VERSION : 0.1
// Data area for commands from master PLC
   VAR
      CRNT_MODE : Int := 1;   // 1 = Auto, 2 = Man, 3 = FatAuto, 4 = FatMan
      HEART_BEAT : Bool;   // Heartbeat
      ESTOP_OK : Bool;   // 1 = OK, 0 = Estop active
      RST_AUT_SEQ : Bool;   // Reset automatic sequence
      RUN_E131 : Bool;   // IA Compressor demand
      RUN_P301 : Bool;   // 1 = Run, 0 = Not
      RUN_BC_SEQ : Bool;   // 1 = Start command. 0 = Not
      PB_STS_CNFMD : Bool;   // Pilot burn status confirmed by IGG
      CRG_BLNK_MODE : Bool;   // 1 = Cargon blanketing mode, 0 = Not
      RUN_BC_O2_RAMP : Bool;   // 1 = Run ramp, 0 = Not
      BC_SD_CMND : Bool;   // 1 = Run. 0 = Shutdown
      STOP_BURNS_CMND : Bool;   // 1 = Burners off, 0 = Not
      CLS_CV127_CMND : Bool;   // 1 = OPEN, 0 = Close
      CLS_CV203_CMND : Bool;   // 1 = Close, 0 = Not
      CLS_CV111_CMND : Bool;   // 1 = Close, 0 = Not
      IGG_ALARM : Bool;   // 1 = IGG Alarm state, 0 = Not
      RUN_P305 : Bool;   // Fresh water pump demand
      CV403_OPEN : Bool;   // 1 = Valve is open, 0 = Not
      "E 500A RUN" : Bool;   // Fuel Pump 1 Enabled
      "E 500B RUN" : Bool;   // Fuel Pump 2 Enabled
      "TIT 360 Healthy" : Bool;   // Outlet CSW Temp TIT360
      "TIT 401 Healthy" : Bool;   // IG Temp
      "PIT 316 Healthy" : Bool;   // Outlet CSW Pressure
      RST_LOCKOUT : Bool;   // Reset alarms
      "CA Blower Running" : Bool;   // E139-MCCP/6TA1
      Alarm_Reset : Bool;   // Alarm_Reset
      BWT_MODE : Bool;
      "P301 PRSNT" : Bool;
      "TIT 315 Healthy" : Bool;   // PIT 315 Healthy
      SFTY_SYS_IL : Bool;   // SFTY_SYS_IL
      "Master Stop" : Bool;   // Master Stop
      "CV401 Closed" : Bool;   // CV401 Closed
      SPR_5_7 : Bool;   // Spare bool
      IGG_CRNT_STEP : Int;   // IGG Current Step
   END_VAR
BEGIN
END_DATA_BLOCK

DATA_BLOCK "55_STATUS_DATA"   // DB55
TITLE = Status Data
{ S7_Optimized_Access := 'FALSE' }
AUTHOR : JRS
VERSION : 0.1
// Data area for status to master PLC
   VAR
      PIT112_SCALED : Real;   // IA Inlet pressure
      CV203_CNTRL : Real;   // Main fuel reg Valve Control
      PIT204_SCALED : Real;   // IGG Inlet fuel pressure
      CRNT_MODE : Int := 1;   // 1 = Auto, 2 = Man, 3 = FatAuto, 4 = FatMan
      HEART_BEAT : Bool;   // Heartbeat
      AUT_SEQ_RNG : Bool;   // Auto sequence running
      VLVS_AT_INIT : Bool;   // All valves in initial state
      P301_ENBLD : Bool;   // P301 enabled input sent from BC
      P301_TRIPPED : Bool;   // P301 tripped input sent from BC
      TS006_OK : Bool;   // TS006 Is healthy
      TS403_OK : Bool;   // TS403 Is healthy
      LS001_OK : Bool;   // LS001 Is healthy
      E131_RUNNING : Bool;   // E131 Running
      BC_SEQ_STARTED : Bool;   // BC Sequence confirmed as started
      PILOT_BURNER_ACTV : Bool;   // Pilot burn confirmed as active
      PILOT_PURGE_DN : Bool;   // Pilot burner purge completed
      RAMPING_O2_ACTV : Bool;   // Ramping of O2 is active
      O2_LVL_OK : Bool;   // O2 Level within specification
      SHTNG_DN_CNF : Bool;   // Shutting down confirmed
      O2_CNTRL_STPD : Bool;   // O2 Control modulation stopped
      BURNS_STOPPED : Bool;   // Confirmation burners are off
      CV127_CLOSED : Bool;   // CV127 Closed status
      CV203_CLOSED : Bool;   // CV203 Closed status
      CV111_CLOSED : Bool;   // CV111 Closed status
      BC_SD_DONE : Bool;   // BC Shutdown sequence done
      BC_ALARM : Bool;   // 1 = BC Alarm state, 0 = Not
      MAA_PRES_IN_RNG : Bool;   // PIT113 Main atom air pressure within range
      "FD001FDU Healthy" : Bool;   // FDU Healthy
      "FS 317 Healthy" : Bool;   // Jacket Cooling Water Flow Switch
      "PIT 204 Healthy" : Bool;   // PIT 204 Healthy
      "FS 320 Healthy" : Bool;   // FS 320 Healthy
      Warnings : Bool;   // Warnings
      "PIT 112 Healthy" : Bool;   // PIT 112 Healthy
      MAIN_BURNER_ACTV : Bool;   // MAIN_BURNER_ACTV
      "BC New ALARM" : Bool;   // New alarm
      "BC New WARNING" : Bool;   // New warning
      P305_ENBLD : Bool;   // P305 enabled input sent from BC
      P305_TRIPPED : Bool;   // P305 tripped input sent from BC
      P305_PRSNT : Bool;   // P305_PRSNT
      SPR_18_3 : Bool;   // Spare bit
      SPR_18_4 : Bool;   // Spare bit
      SPR_18_5 : Bool;   // Spare bit
      SPR_18_6 : Bool;   // Spare bit
      SPR_18_7 : Bool;   // Spare bit
   END_VAR
BEGIN
END_DATA_BLOCK

DATA_BLOCK "57_COMMS_DATE_TIME"   // DB57
{ S7_Optimized_Access := 'FALSE' }
VERSION : 0.1
   VAR
      SYSTEM_TIME : DTL;
      LOCAL_TIME : DTL;
   END_VAR
BEGIN
END_DATA_BLOCK

DATA_BLOCK "59_COMMS_HEALTH_DATA"   // DB59
TITLE = Communications Health Data
{ S7_Optimized_Access := 'TRUE' }
AUTHOR : JRS
VERSION : 0.1
// Data area for communications health determination
   VAR
      CLOCK_POS_EDGE : Bool;   // Edge bit
      CLOCK_NEG_EDGE : Bool;   // Edge bit
      MSTR_TRUE_TMR : TON_TIME;
      MSTR_FALSE_TMR : TON_TIME;
      MSTR_HB_MISSING : Bool;   // Heatbeat missing flag
   END_VAR
BEGIN
   MSTR_FALSE_TMR.PT := T#2s;
   MSTR_TRUE_TMR.PT := T#2s;
END_DATA_BLOCK

// folder: 60 - 69 Alarm & Satus Handling

DATA_BLOCK "60_Alarm_Data"   // DB60
{ S7_Optimized_Access := 'FALSE' }
VERSION : 0.1
   VAR
      BC_ALARM_WORD_01 : Word;
      BC_ALARM_WORD_02 : Word;
      BC_ALARM_WORD_03 : Word;
      BC_ALARM_WORD_04 : Word;
      BC_ALARM_WORD_05 : Word;
      BC_ALARM_WORD_06 : Word;
      BC_ALARM_WORD_07 : Word;
      BC_ALARM_WORD_08 : Word;
      BC_ALARM_WORD_09 : Word;
      BC_ALARM_WORD_10 : Word;
      BC_ALARM_WORD_11 : Word;
      BC_ALARM_WORD_12 : Word;
      BC_ALARM_WORD_13 : Word;
      BC_ALARM_WORD_14 : Word;
      BC_ALARM_WORD_15 : Word;
      BC_ALARM_WORD_16 : Word;
      ALRM_PRSNT : Bool;
   END_VAR
BEGIN
END_DATA_BLOCK

DATA_BLOCK "62_Warning_Data"   // DB62
{ S7_Optimized_Access := 'FALSE' }
VERSION : 0.1
   VAR
      BC_WARNING_WORD_01 : Word;   // PIT 204
      BC_WARNING_WORD_02 : Word;   // TIT 202
      BC_WARNING_WORD_03 : Word;   // PIT 205
      BC_WARNING_WORD_04 : Word;   // PIT 112
      BC_WARNING_WORD_05 : Word;   // PIT 113
      BC_WARNING_WORD_06 : Word;
      BC_WARNING_WORD_07 : Word;
      BC_WARNING_WORD_08 : Word;
      WRNG_PRSNT : Bool;
   END_VAR
BEGIN
END_DATA_BLOCK

DATA_BLOCK "503_WARNING CHCK_DB"   // DB63
{ S7_Optimized_Access := 'TRUE' }
VERSION : 0.1
// stored: InstanceOfName 503_ALARM CHCK
"503_ALARM CHCK"
BEGIN
END_DATA_BLOCK

DATA_BLOCK "64_Message_Data"   // DB64
{ S7_Optimized_Access := 'FALSE' }
VERSION : 0.1
   VAR
      BC_MESSAGE_WORD_01 : Word;
      BC_MESSAGE_WORD_02 : Word;
      BC_MESSAGE_WORD_03 : Word;
      BC_MESSAGE_WORD_04 : Word;
      BC_MESSAGE_WORD_05 : Word;
      BC_MESSAGE_WORD_06 : Word;
      BC_MESSAGE_WORD_07 : Word;
      BC_MESSAGE_WORD_08 : Word;
      MSG_PRSNT : Bool;
   END_VAR
BEGIN
END_DATA_BLOCK

DATA_BLOCK "503_ALARM CHCK_DB"   // DB65
{ S7_Optimized_Access := 'TRUE' }
VERSION : 0.1
// stored: InstanceOfName 503_ALARM CHCK
"503_ALARM CHCK"
BEGIN
END_DATA_BLOCK

DATA_BLOCK "66_Event_Data"   // DB66
{ S7_Optimized_Access := 'FALSE' }
VERSION : 0.1
   VAR
      BC_EVENT_WORD_01 : Word;
      BC_EVENT_WORD_02 : Word;
      BC_EVENT_WORD_03 : Word;
      BC_EVENT_WORD_04 : Word;
      BC_EVENT_WORD_05 : Word;
      BC_EVENT_WORD_06 : Word;
      BC_EVENT_WORD_07 : Word;
      BC_EVENT_WORD_08 : Word;
      EVENT_PRSNT : Bool;
   END_VAR
BEGIN
END_DATA_BLOCK

DATA_BLOCK "68_Sys_Status_Data"   // DB68
TITLE = System Status Data
{ S7_Optimized_Access := 'TRUE' }
AUTHOR : JRS
VERSION : 0.1
// Data area for system status information as required by the code
   VAR
      VLVS_AT_INIT : Bool;   // All valves at initial position
      INTRLKS_OK : Bool;   // System interlocks ok
      IA_PRES_IN_RNG : Bool;   // IA Pressure Within Range - PIT112
      CSW_IL_PRES_IN_RNG : Bool;   // CSW Inlet pressure within range - PIT359
      FUEL_PRES_IN_RNG : Bool;   // Fuel pressure within range - PIT204
      OP_PRES_IN_RNG : Bool;   // Output pressure within range - PIT402
      VALID_FLAME : Bool;   // Flame detection & > min value - FD001
      O2_INTO_SPEC_DLY : TON_TIME;   // O2 Going into specification de-bounce timer
      O2_OUT_SPEC_DLY : TOF_TIME;   // O2 Going out of specification de-bounce timer
      O2_WITHIN_SPEC : Bool;   // O2 Contenct is within specification
      SHT_DN_CNF_DLY : TP_TIME;   // Shutting down confirmed timer
      O2_CNTRL_STPPD_DLY : TP_TIME;   // O2 Control stopped confirmed timer
      BURNS_STPPD_DLY : TP_TIME;   // Burns stopped confirmed timer
      CV127_CLSD_DLY : TP_TIME;   // CV127 Closed confirmed timer
      CV203_CLSD_DLY : TON_TIME;   // CV203 Closed confirmed timer
      CV111_CLSD_DLY : TON_TIME;   // CV111 Closed confirmed timer
      BC_SD_DONE : TP_TIME;   // BC Shutdown done timer
      CV127_CLSD_FLG : Bool;
   END_VAR
BEGIN
END_DATA_BLOCK

DATA_BLOCK "Main Burner Animation_DB"   // DB69
{ S7_Optimized_Access := 'TRUE' }
VERSION : 0.1
// stored: InstanceOfName Animation
"Animation"
BEGIN
END_DATA_BLOCK

DATA_BLOCK "IDB_E131_Animation"   // DB132
{ S7_Optimized_Access := 'TRUE' }
VERSION : 0.1
// stored: InstanceOfName Animation
"Animation"
BEGIN
END_DATA_BLOCK

DATA_BLOCK "64_Functioning Hours_P301_IDB"   // DB301
{ S7_Optimized_Access := 'TRUE' }
VERSION : 0.1
// stored: InstanceOfName 64_Functioning Hours
"64_Functioning Hours"
BEGIN
END_DATA_BLOCK

DATA_BLOCK "Animation_P301_IDB"   // DB302
{ S7_Optimized_Access := 'TRUE' }
VERSION : 0.1
// stored: InstanceOfName Animation
"Animation"
BEGIN
END_DATA_BLOCK

DATA_BLOCK "IDB_E-600"   // DB600
{ S7_Optimized_Access := 'FALSE' }
VERSION : 0.1
// stored: InstanceOfName 502_ALM_ANALOG
"502_ALM_ANALOG"
BEGIN
END_DATA_BLOCK

DATA_BLOCK "IDB_E700 Alarms"   // DB701
{ S7_Optimized_Access := 'FALSE' }
VERSION : 0.1
// stored: InstanceOfName 502_ALM_ANALOG
"502_ALM_ANALOG"
BEGIN
END_DATA_BLOCK

DATA_BLOCK "P305_Functioning Hours_IDB"   // DB705
{ S7_Optimized_Access := 'TRUE' }
VERSION : 0.1
// stored: InstanceOfName 64_Functioning Hours
"64_Functioning Hours"
BEGIN
END_DATA_BLOCK

DATA_BLOCK "P305_Animation_IDB"   // DB706
{ S7_Optimized_Access := 'TRUE' }
VERSION : 0.1
// stored: InstanceOfName Animation
"Animation"
BEGIN
END_DATA_BLOCK

DATA_BLOCK "IDB_PIT 112"   // DB712
{ S7_Optimized_Access := 'FALSE' }
VERSION : 0.1
// stored: InstanceOfName 502_ALM_ANALOG
"502_ALM_ANALOG"
BEGIN
END_DATA_BLOCK

DATA_BLOCK "IDB_PIT 113"   // DB713
{ S7_Optimized_Access := 'FALSE' }
VERSION : 0.1
// stored: InstanceOfName 502_ALM_ANALOG
"502_ALM_ANALOG"
BEGIN
END_DATA_BLOCK

DATA_BLOCK "IDB_FD-001"   // DB721
{ S7_Optimized_Access := 'FALSE' }
VERSION : 0.1
// stored: InstanceOfName 502_ALM_ANALOG
"502_ALM_ANALOG"
BEGIN
END_DATA_BLOCK

DATA_BLOCK "IDB_TIT 202"   // DB722
{ S7_Optimized_Access := 'FALSE' }
VERSION : 0.1
// stored: InstanceOfName 502_ALM_ANALOG
"502_ALM_ANALOG"
BEGIN
END_DATA_BLOCK

DATA_BLOCK "IDB_PIT 204"   // DB724
{ S7_Optimized_Access := 'FALSE' }
VERSION : 0.1
// stored: InstanceOfName 502_ALM_ANALOG
"502_ALM_ANALOG"
BEGIN
END_DATA_BLOCK

DATA_BLOCK "IDB_PIT 205"   // DB725
{ S7_Optimized_Access := 'FALSE' }
VERSION : 0.1
// stored: InstanceOfName 502_ALM_ANALOG
"502_ALM_ANALOG"
BEGIN
END_DATA_BLOCK

// folder: 70 - 79 Modes of Operation

DATA_BLOCK "70_Mode_Data"   // DB70
{ S7_Optimized_Access := 'TRUE' }
VERSION : 0.1
   VAR
      CRNT_MODE : Int := 1;   // 1 = Auto, 2 = Man, 3 = FatAuto, 4 = FatMan
      INTO_AUTO : Bool;   // Transition to auto
      IN_MAN : Bool;   // In manual
      INTO_AUT_PLS : Bool;   // Pulse bit
      AUT_RST_PLS : TP_TIME;   // Automatic sequence reset pulse
   END_VAR
BEGIN
   AUT_RST_PLS.PT := T#1s;
END_DATA_BLOCK

// folder: 80 - 89 HMI Handling

DATA_BLOCK "80_From_HMI"   // DB80
{ S7_Optimized_Access := 'TRUE' }
VERSION : 0.1
   VAR
      FAT_Mode : Bool := False;   // Set or Reset in HMI
      RST_AUT_SEQ : Bool;   // Reset automatic sequence
      IGG_STND_ALN : Bool := 0;   // 0 = Part of BWT, 1 = Stand Alone
   END_VAR
   VAR RETAIN
      BWT_BYPASS : Bool := FALSE;   // 0 = BWT Control, 1 = BWT Bypassed
      P301_PRSNT : Bool := TRUE;   // 1 = CSW Pump fitted, 0 = Not
      CV312_PRSNT : Bool := FALSE;   // 1 = Scrubber valve fitted, 0 = Not
   END_VAR
   VAR
      MAN_DQ_0_0 : Bool;   // Q0.0 - Test Pressure Valve Control (CV-127)
      MAN_DQ_0_1 : Bool;   // Q0.1 - Pilot B Ignition Air Valve Control (CV-124)
      MAN_DQ_0_2 : Bool;   // Q0.2 - Pilot B Fuel Valve 1 Control (CV-215)
      MAN_DQ_0_3 : Bool;   // Q0.3 - Pilot B Fuel Valve 2 Control (CV-216)
      MAN_DQ_0_4 : Bool;   // Q0.4 - Main B Atom Air Valve Control (CV-114)
      MAN_DQ_0_5 : Bool;   // Q0.5 - Main B Fuel Valve 1 Control (CV-206)
      MAN_DQ_0_6 : Bool;   // Q0.6 - Main B Fuel Valve 2 Control (CV-207)
      MAN_DQ_0_7 : Bool;   // Q0.7 - IA Comp Control (E131)
      MAN_DQ_1_0 : Bool;   // Q1.0 - CSW Pump Control (P301)
      MAN_DQ_1_1 : Bool;   // Q1.1 - Igniter Control (X-001)
      MAN_DQ_1_2 : Bool;   // Q1.2 - Spare output
      MAN_DQ_1_3 : Bool;   // Q1.3 - Spare output
      MAN_DQ_1_4 : Bool;   // Q1.4 - Spare output
      MAN_DQ_1_5 : Bool;   // Q1.5 - Spare output
      MAN_DQ_1_6 : Bool;   // Q1.6 - Spare output
      MAN_DQ_1_7 : Bool;   // Q1.7 - Fresh Water Pump Control (P-305)
      MAN_AQ_INC_96 : Bool;   // QW96 - Spare - Increase % Signal
      MAN_AQ_DEC_96 : Bool;   // QW96 - Spare - Decrease % Signal
      MAN_AQ_INC_98 : Bool;   // QW96 - Spare - Increase % Signal
      MAN_AQ_DEC_98 : Bool;   // QW96 - Spare - Decrease % Signal
      MAN_AQ_INC_100 : Bool;   // QW100 - CV203 - Increase % Signal
      MAN_AQ_DEC_100 : Bool;   // QW100 - CV203 - Decrease % Signal
      MAN_AQ_INC_102 : Bool;   // QW102 - CV111 - Increase % Signal
      MAN_AQ_DEC_102 : Bool;   // QW102 - CV111 - Decrease % Signal
      FLM_FAIL_DLY : Time := T#1s;   // Flame fail delay
      "Reset CV203 PID" : Bool;
   END_VAR
   VAR RETAIN
      BurnerProgramedStop : Bool := false;
      P305_PRSNT : Bool := TRUE;
   END_VAR
BEGIN
END_DATA_BLOCK

DATA_BLOCK "82_To_HMI"   // DB82
{ S7_Optimized_Access := 'TRUE' }
VERSION : 0.1
   VAR
      CRNT_MODE : Int := 1;   // 1 = Man, 2 = Auto, 3 = FAT Man, 4 = FATAuto
      "Test Fuel Control" : Real;
   END_VAR
   VAR RETAIN
      "I&A Compressor Run Days" : Int;
      "I&A Compressor Run Hours" : Int;
      "I&A Compressor Run Minutes" : Int;
      "I&A Compressor Run Seconds" : Int;
   END_VAR
   VAR
      "I&A Compressor Reset Hours" : Bool;
   END_VAR
   VAR RETAIN
      "I&A Compressor Total Run Hours" : Int;
   END_VAR
   VAR
      "I&A Compressor Service Due" : Bool;
   END_VAR
   VAR RETAIN
      "I&A Compressor Service Time Hours" : Int;
      "I&A Compressor Service Time Days" : Int;
      "I&A Compressor Hours to Service" : Int;
   END_VAR
   VAR
      "IA Compressor Animation" : Int;
   END_VAR
   VAR RETAIN
      "P301 CSW Pump Run Days" : Int;
      "P301 CSW Pump Run Hours" : Int;
      "P301 CSW Pump Run Minutes" : Int;
      "P301 CSW Pump Run Seconds" : Int;
   END_VAR
   VAR
      "P301 CSW Pump Reset Hours" : Bool;
   END_VAR
   VAR RETAIN
      "P301 CSW Pump Total Run Hours" : Int;
   END_VAR
   VAR
      "P301 CSW Pump Service Due" : Bool;
   END_VAR
   VAR RETAIN
      "P301 CSW Pump Service Time Hours" : Int;
      "P301 CSW Pump Service Time Days" : Int;
      "P301 CSW Pump Hours to Service" : Int;
   END_VAR
   VAR
      "P301 CSW Pump Animation" : Int;
      "P305 FW Pump Run Days" : Int;
      "P305 FW Pump Run Hours" : Int;
      "P305 FW Pump Run Minutes" : Int;
      "P305 FW Pump Run Seconds" : Int;
      "P305 FW Pump Reset Hours" : Bool;
      "P305 FW Pump Total Run Hours" : Int;
      "P305 FW Pump Service Due" : Bool;
      "P305 FW Pump Service Time Hours" : Int;
      "P305 FW Pump Service Time Days" : Int;
      "P305 FW Pump Hours to Service" : Int;
      "P305 FW Pump Animation" : Int;
      "E-STOP LATCHED" : Bool;
   END_VAR
BEGIN
END_DATA_BLOCK

DATA_BLOCK "84_Setpoints"   // DB84
{ S7_Optimized_Access := 'TRUE' }
VERSION : 0.1
   VAR RETAIN
      FD001_Min : Real := 30.0;   // FD001 sensor pilot target setpoint
      FD001_LowLow : Real := 30.0;   // FD001 sensor pilot low low setpoint
      FD001_Low : Real := 40.0;   // FD001 sensor pilot low setpoint
      PIT113_Pilot_Target : Real := 7.0;   // PIT113 sensor target setpoint (bar g)
   END_VAR
   VAR
      PIT113_Burner_Target : Real := 7.0;
   END_VAR
   VAR RETAIN
      PIT113_LowLow : Real := 2.5;   // PIT113 sensor low low setpoint (bar g)
      PIT113_Low : Real := 3.0;   // PIT113 sensor low setpoint (bar g)
      PIT113_High : Real := 12.0;   // PIT113 sensor high setpoint (bar g)
      PIT113_HighHigh : Real := 13.0;   // PIT113 sensor high high setpoint (bar g)
      PIT205_Target : Real := 6.89;   // PIT205 sensor target setpoint (bar g)
      PIT205_LowLow : Real := 0.8;   // PIT205 sensor low low setpoint (bar g)
      PIT205_Low : Real := 0.9;   // PIT205 sensor low setpoint (bar g)
      PIT205_High : Real := 12.0;   // PIT205 sensor high setpoint (bar g)
      PIT205_HighHigh : Real := 12.5;   // PIT205 sensor high high setpoint (bar g)
      TIT202_LowLow : Real := 3.0;   // TIT202 sensor low low setpoint (degC)
      TIT202_Low : Real := 4.0;   // TIT202 sensor low setpoint (degC)
      TIT202_High : Real := 50.0;   // TIT202 sensor high setpoint (degC)
      TIT202_HighHigh : Real := 55.0;   // TIT202 sensor high high setpoint (degC)
      E600_BWT_LowLow : Real := 0.0;   // TX600 sensor ballast water treatment mode low low setpoint (%)
      E600_BWT_Low : Real := 0.05;   // TX600 sensor ballast water treatment mode low setpoint (%)
      E600_BWT_Target : Real := 0.2;   // TX600 sensor balast water treatment mode target setpoint (%)
      E600_BWT_High : Real := 0.5;   // TX600 sensor ballast water treatment mode high setpoint (%)
      E600_BWT_HighHigh : Real := 0.6;   // TX600 sensor ballast water treatment mode high high setpoint (%)
      E600_CB_LowLow : Real := 2.0;   // TX600 sensor cargo blanketing mode low low setpoint (%)
      E600_CB_Low : Real := 2.5;   // TX600 sensor cargo blanketing mode low setpoint (%)
      E600_CB_Target : Real := 3.0;   // TX600 sensor cargo blanketing mode target setpoint (%)
      E600_CB_High : Real := 4.0;   // TX600 sensor cargo blanketing mode high setpoint (%)
      E600_CB_HighHigh : Real := 4.5;   // TX600 sensor cargo blanketing mode high high setpoint (%)
      TX700_Low : Real := 0.0;   // TX700 sensor low setpoint (ppm)
      TX700_High : Real := 30.0;   // TX700 sensor high setpoint (ppm)
      PIT204_Target : Real := 5.0;   // PIT204 sensor target setpoint (bar g)
      PIT204_LowLow : Real := 0.5;   // PIT204 sensor low low setpoint (bar g)
      PIT204_Low : Real := 0.6;   // PIT204 sensor low setpoint (bar g)
      PIT204_High : Real := 12.0;   // PIT204 sensor high setpoint (bar g)
      PIT204_HighHigh : Real := 12.5;   // PIT204 sensor high high setpoint (bar g)
      PIT112_Target : Real := 7.5;   // PIT112 sensor target setpoint (bar g)
      PIT112_LowLow : Real := 2.5;   // PIT112 sensor low low setpoint (bar g)
      PIT112_Low : Real := 3.0;   // PIT112 sensor low setpoint (bar g)
      PIT112_High : Real := 12.0;   // PIT112 sensor high setpoint (bar g)
      PIT112_HighHigh : Real := 13.0;   // PIT112 sensor high high setpoint (bar g)
      P_ON : Bool := FALSE;
      I_ON : Bool := TRUE;
      D_ON : Bool := TRUE;
      Gain : Real := 0.005;
      "Integration Time" : Time := T#1S_950MS;
      "Derive Time" : Time := T#100MS;
      "Max Opening" : Real := 80.0;
      "Min Opening" : Real := 55.0;
   END_VAR
BEGIN
END_DATA_BLOCK

DATA_BLOCK "86_Times"   // DB86
{ S7_Optimized_Access := 'TRUE' }
VERSION : 0.1
   VAR
      "CV127_OPEN_TIME_#1" : Time := T#2S;   // CV127 Open Delay #1
      CV127_CLOSED_TIME : Time := T#2S;   // CV127 Closed Delay
      "CV127_OPEN_TIME_#2" : Time := T#2S;   // CV127 Open Delay #2
      CV124_OPEN_TIME : Time := T#2S;   // CV124 Open Delay
      CV124_CLOSE_TIME_PRG : Time := T#2S;   // CV124 Close Delay Purging
      CV114_OPEN_TIME : Time := T#2S;   // CV114 Open Delay
      CV206_OPEN_TIME : Time := T#2S;   // CV206 Open Delay
      CV207_OPEN_TIME : Time := T#2S;   // CV207 Open Delay
      CV215_OPEN_TIME : Time := T#2S;   // CV215 Open Delay
      CV215_CLOSE_TIME_PRG : Time := T#2S;   // CV215 Close Delay Purging
      CV216_OPEN_TIME : Time := T#2S;   // CV216 Open Delay
      CV216_CLOSE_TIME_PRG : Time := T#2S;   // CV216 Close Delay Purging
      CV216_OPEN_TIME_PRG : Time := T#2S;   // CV216 Open Delay Purging
      CV206_CLOSE_TIME : Time := T#2S;   // CV206 Close Delay
      CV207_CLOSE_TIME : Time := T#2S;   // CV207 Close Delay
      CV114_CLOSE_TIME : Time := T#2S;   // CV114 Close Delay
      CV215_CLOSE_TIME : Time := T#2S;   // CV215 Close Delay
      CV216_CLOSE_TIME : Time := T#2S;   // CV216 Close Delay
      CV124_CLOSE_TIME : Time := T#2S;   // CV124 Close Delay
      X001_MAX_RUN_TIME : Time := T#5S;   // X001 Max continuous run time of igniter
      X001_RUN_CNF_TIME : Time := T#3S;   // X001 Run confirmation time
      FD_DET_DELAY : Time := T#3S;   // Flame detection delay
      FD_VRFCTN_TIME : Time := T#5S;   // Flame verification time
      FDU_DET_TIME : Time := T#5S;   // FDU Flame detection time
      MAX_IGNTN_SEQ_TIME : Time := T#1M;   // Maximum ignition sequence run time
      MAX_MAIN_BURN_SEQ_TIME : Time := T#1H;   // Maximum main burner sequence run time
      MAX_PILOT_PURGE_SEQ_TIME : Time := T#30S;   // Maximum pilot burner purge sequence run time
      O2_CHECK_TIME : Time := T#20S;   // Time for O2 check after valve change
      STEP_MAX_TIME_STP_001 : Time := T#30MS;
      STEP_MAX_TIME_STP_005 : Time := T#30MS;
      STEP_MAX_TIME_STP_010 : Time := T#30MS;
      STEP_MAX_TIME_STP_020 : Time := T#30MS;
      STEP_MAX_TIME_STP_025 : Time := T#30MS;
      STEP_MAX_TIME_STP_027 : Time := T#30MS;
      STEP_MAX_TIME_STP_029 : Time := T#30MS;
      STEP_MAX_TIME_STP_030 : Time := T#30MS;
      STEP_MAX_TIME_STP_040 : Time := T#30MS;
      STEP_MAX_TIME_STP_050 : Time := T#30MS;
      STEP_MAX_TIME_STP_060 : Time := T#30MS;
      STEP_MAX_TIME_STP_070 : Time := T#30MS;
      STEP_MAX_TIME_STP_080 : Time := T#30MS;
      STEP_MAX_TIME_STP_090 : Time := T#30MS;
      STEP_MAX_TIME_STP_095 : Time := T#30MS;
      STEP_MAX_TIME_STP_100 : Time := T#30MS;
      STEP_MAX_TIME_STP_110 : Time := T#30MS;
      STEP_MAX_TIME_STP_120 : Time := T#30MS;
      STEP_MAX_TIME_STP_130 : Time := T#30MS;
      STEP_MAX_TIME_STP_140 : Time := T#30MS;
      STEP_MAX_TIME_STP_150 : Time := T#30MS;
      STEP_MAX_TIME_STP_160 : Time := T#1M_100MS;
      STEP_MAX_TIME_STP_170 : Time := T#30MS;
      STEP_MAX_TIME_STP_180 : Time := T#30MS;
      STEP_MAX_TIME_STP_190 : Time := T#30MS;
      STEP_MAX_TIME_STP_200 : Time := T#30MS;
      STEP_MAX_TIME_STP_210 : Time := T#30MS;
      STEP_MAX_TIME_STP_220 : Time := T#30MS;
      STEP_MAX_TIME_STP_230 : Time := T#30MS;
      STEP_MAX_TIME_STP_240 : Time := T#30MS;
      STEP_MAX_TIME_STP_250 : Time := T#30MS;
      STEP_MAX_TIME_STP_260 : Time := T#30MS;
      STEP_MAX_TIME_STP_270 : Time := T#30MS;
      STEP_MAX_TIME_STP_280 : Time := T#30MS;
      STEP_MAX_TIME_STP_290 : Time := T#30MS;
      STEP_MAX_TIME_STP_300 : Time := T#30MS;
      STEP_MAX_TIME_STP_310 : Time := T#30MS;
      STEP_MAX_TIME_STP_320 : Time := T#30MS;
      STEP_MAX_TIME_STP_330 : Time := T#30MS;
      STEP_MAX_TIME_STP_340 : Time := T#30MS;
      STEP_MAX_TIME_STP_350 : Time := T#30MS;
      STEP_MAX_TIME_STP_360 : Time := T#30MS;
      STEP_MAX_TIME_STP_370 : Time := T#30MS;
      STEP_MAX_TIME_STP_380 : Time := T#30MS;
      STEP_MAX_TIME_STP_390 : Time := T#30MS;
      STEP_MAX_TIME_STP_400 : Time := T#30MS;
      STEP_MAX_TIME_STP_410 : Time := T#30MS;
      STEP_MAX_TIME_STP_420 : Time := T#30MS;
      STEP_MAX_TIME_STP_430 : Time := T#30MS;
      STEP_MAX_TIME_STP_440 : Time := T#30MS;
      STEP_MAX_TIME_STP_450 : Time := T#30MS;
      STEP_MAX_TIME_STP_460 : Time := T#30MS;
      STEP_MAX_TIME_STP_470 : Time := T#30MS;
      STEP_MAX_TIME_STP_480 : Time := T#30MS;
      STEP_MAX_TIME_STP_490 : Time := T#30MS;
      STEP_MAX_TIME_STP_500 : Time := T#30MS;
      STEP_MAX_TIME_STP_510 : Time := T#30MS;
      STEP_MAX_TIME_STP_520 : Time := T#30MS;
      STEP_MAX_TIME_STP_525 : Time := T#30MS;
      STEP_MAX_TIME_STP_530 : Time := T#30MS;
      STEP_MAX_TIME_STP_540 : Time := T#30MS;
      STEP_MAX_TIME_STP_550 : Time := T#30MS;
      STEP_MAX_TIME_STP_560 : Time := T#30MS;
      STEP_MAX_TIME_STP_570 : Time := T#30MS;
   END_VAR
   VAR RETAIN
      "FS317 delay" : Time := T#5S;
      "FS320 delay" : Time := T#5S;
   END_VAR
   VAR
      "PS101 Alarm Delay" : Time := T#1M;
   END_VAR
BEGIN
END_DATA_BLOCK

// folder: 90 - 99 Manual Functions

DATA_BLOCK "90_Manual_Data"   // DB90
{ S7_Optimized_Access := 'TRUE' }
VERSION : 0.1
   VAR
      INC_PLS_96 : Bool;   // Pulse bit
      INC_PLS_96_Hz : Bool;   // Pulse bit
      DEC_PLS_96 : Bool;   // Pulse bit
      DEC_PLS_96_Hz : Bool;   // Pulse bit
      INC_PLS_98 : Bool;   // Pulse bit
      INC_PLS_98_Hz : Bool;   // Pulse bit
      DEC_PLS_98 : Bool;   // Pulse bit
      DEC_PLS_98_Hz : Bool;   // Pulse bit
      INC_PLS_100 : Bool;   // Pulse bit
      INC_PLS_100_Hz : Bool;   // Pulse bit
      DEC_PLS_100 : Bool;   // Pulse bit
      DEC_PLS_100_Hz : Bool;   // Pulse bit
      INC_PLS_102 : Bool;   // Pulse bit
      INC_PLS_102_Hz : Bool;   // Pulse bit
      DEC_PLS_102 : Bool;   // Pulse bit
      DEC_PLS_102_Hz : Bool;   // Pulse bit
   END_VAR
BEGIN
END_DATA_BLOCK

// folder: (top level)

ORGANIZATION_BLOCK "BC Main PLC"   // OB1, LAD, ProgramCycle
TITLE = "Main Program Sweep (Cycle)"
{ S7_Optimized_Access := 'TRUE' }
VERSION : 0.1
   VAR_INPUT
      Initial_Call : Bool;   // Initial call of this OB
      Remanence : Bool;   // =True, if remanent data are available
   END_VAR
   VAR_TEMP   // added for the SCL form of the ladder/FBD networks
      _w1 : Bool;
   END_VAR
BEGIN

REGION Network 1: Digital Input Processing
   // To process raw inputs prior to code use
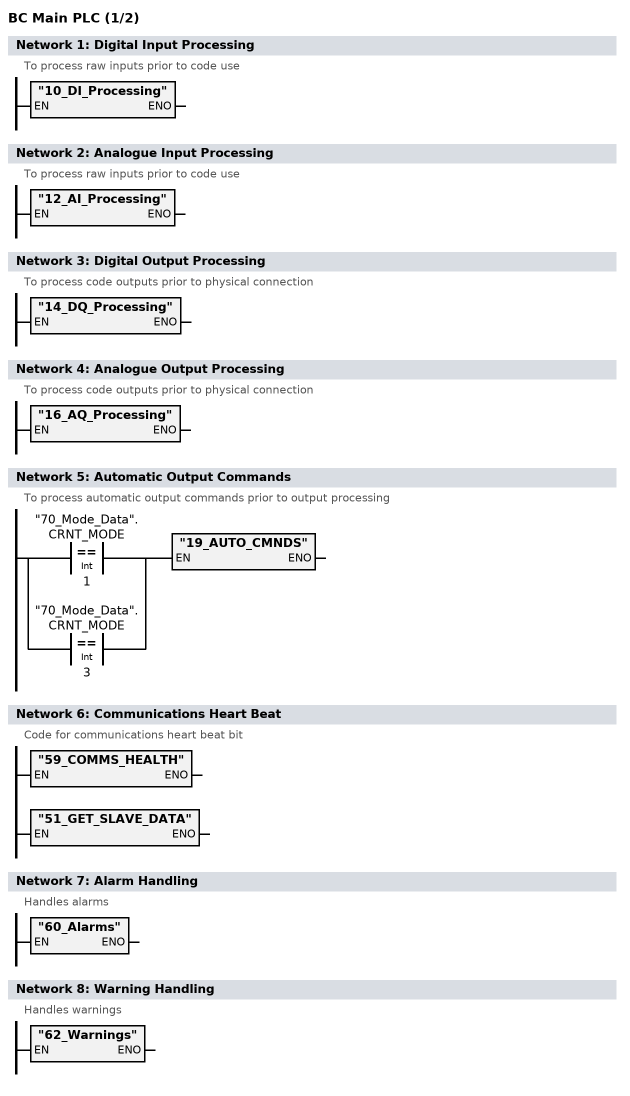
   RUNG wire#powerrail
      "10_DI_Processing"()
   END_RUNG
   // the same network as SCL:
   "10_DI_Processing"();
END_REGION

REGION Network 2: Analogue Input Processing
   // To process raw inputs prior to code use
   RUNG wire#powerrail
      "12_AI_Processing"()
   END_RUNG
   // the same network as SCL:
   "12_AI_Processing"();
END_REGION

REGION Network 3: Digital Output Processing
   // To process code outputs prior to physical connection
   RUNG wire#powerrail
      "14_DQ_Processing"()
   END_RUNG
   // the same network as SCL:
   "14_DQ_Processing"();
END_REGION

REGION Network 4: Analogue Output Processing
   // To process code outputs prior to physical connection
   RUNG wire#powerrail
      "16_AQ_Processing"()
   END_RUNG
   // the same network as SCL:
   "16_AQ_Processing"();
END_REGION

REGION Network 5: Automatic Output Commands
   // To process automatic output commands prior to output processing
   RUNG wire#powerrail
      { S7_Templates := "SrcType := Int" } EQ_Contact(in1 := "70_Mode_Data".CRNT_MODE, in2 := 1)
      wire#w1
      "19_AUTO_CMNDS"()
   END_RUNG
   RUNG wire#powerrail
      { S7_Templates := "SrcType := Int" } EQ_Contact(in1 := "70_Mode_Data".CRNT_MODE, in2 := 3)
   END_RUNG wire#w1
   // the same network as SCL:
   IF ("70_Mode_Data".CRNT_MODE = 1) OR ("70_Mode_Data".CRNT_MODE = 3) THEN "19_AUTO_CMNDS"(); END_IF;
END_REGION

REGION Network 6: Communications Heart Beat
   // Code for communications heart beat bit
   RUNG wire#powerrail
      "59_COMMS_HEALTH"()
   END_RUNG
   RUNG wire#powerrail
      "51_GET_SLAVE_DATA"()
   END_RUNG
   // the same network as SCL:
   "59_COMMS_HEALTH"();
   "51_GET_SLAVE_DATA"();
END_REGION

REGION Network 7: Alarm Handling
   // Handles alarms
   RUNG wire#powerrail
      "60_Alarms"()
   END_RUNG
   // the same network as SCL:
   "60_Alarms"();
END_REGION

REGION Network 8: Warning Handling
   // Handles warnings
   RUNG wire#powerrail
      "62_Warnings"()
   END_RUNG
   // the same network as SCL:
   "62_Warnings"();
END_REGION

REGION Network 9: Message Handling
   // Handles messages
END_REGION

REGION Network 10: Event Handling
   // Record events
END_REGION

REGION Network 11: System Processing
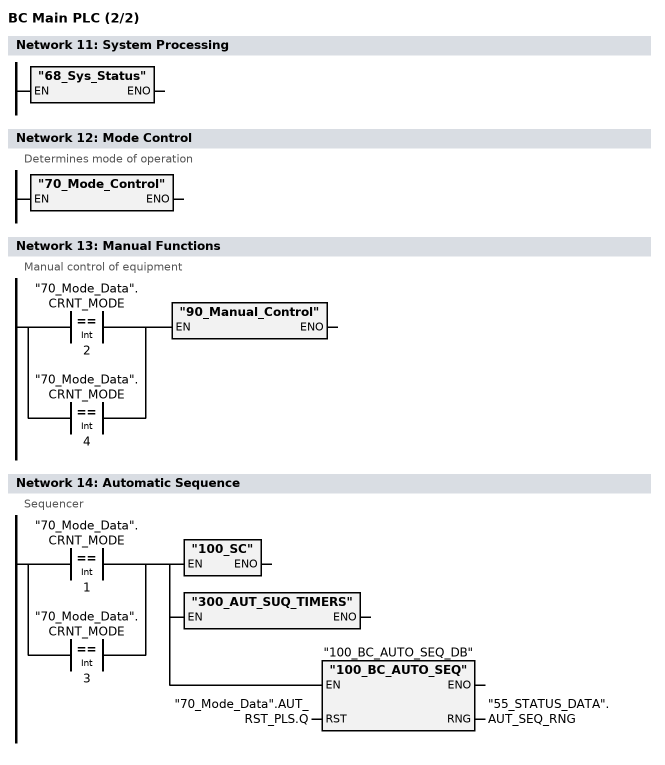
   RUNG wire#powerrail
      "68_Sys_Status"()
   END_RUNG
   // the same network as SCL:
   "68_Sys_Status"();
END_REGION

REGION Network 12: Mode Control
   // Determines mode of operation
   RUNG wire#powerrail
      "70_Mode_Control"()
   END_RUNG
   // the same network as SCL:
   "70_Mode_Control"();
END_REGION

REGION Network 13: Manual Functions
   // Manual control of equipment
   RUNG wire#powerrail
      { S7_Templates := "SrcType := Int" } EQ_Contact(in1 := "70_Mode_Data".CRNT_MODE, in2 := 2)
      wire#w1
      "90_Manual_Control"()
   END_RUNG
   RUNG wire#powerrail
      { S7_Templates := "SrcType := Int" } EQ_Contact(in1 := "70_Mode_Data".CRNT_MODE, in2 := 4)
   END_RUNG wire#w1
   // the same network as SCL:
   IF ("70_Mode_Data".CRNT_MODE = 2) OR ("70_Mode_Data".CRNT_MODE = 4) THEN "90_Manual_Control"(); END_IF;
END_REGION

REGION Network 14: Automatic Sequence
   // Sequencer
   RUNG wire#powerrail
      { S7_Templates := "SrcType := Int" } EQ_Contact(in1 := "70_Mode_Data".CRNT_MODE, in2 := 1)
      wire#w1
      "100_SC"()
   END_RUNG
   RUNG wire#powerrail
      { S7_Templates := "SrcType := Int" } EQ_Contact(in1 := "70_Mode_Data".CRNT_MODE, in2 := 3)
   END_RUNG wire#w1
   RUNG wire#w1
      "300_AUT_SUQ_TIMERS"()
   END_RUNG
   RUNG wire#w1
      "100_BC_AUTO_SEQ_DB"(RST := "70_Mode_Data".AUT_RST_PLS.Q, RNG => "55_STATUS_DATA".AUT_SEQ_RNG)
   END_RUNG
   // the same network as SCL:
   #_w1 := ("70_Mode_Data".CRNT_MODE = 1) OR ("70_Mode_Data".CRNT_MODE = 3);
   IF #_w1 THEN
       "100_SC"();
       "300_AUT_SUQ_TIMERS"();
       "100_BC_AUTO_SEQ_DB"(RST := "70_Mode_Data".AUT_RST_PLS.Q, RNG => "55_STATUS_DATA".AUT_SEQ_RNG);   // "100_BC_AUTO_SEQ"
   END_IF;
END_REGION
END_ORGANIZATION_BLOCK

// folder: 10 - 19 IO & Processing

FUNCTION "10_DI_Processing" : Void   // FC10, LAD
TITLE = Digital Input Processing
{ S7_Optimized_Access := 'TRUE' }
AUTHOR : JRS
VERSION : 0.1
// To process raw inputs prior to code use
BEGIN

REGION Network 1: I0.0 - CA Pressure Switch OK (PS-101)
   // True = OK, False = NOK
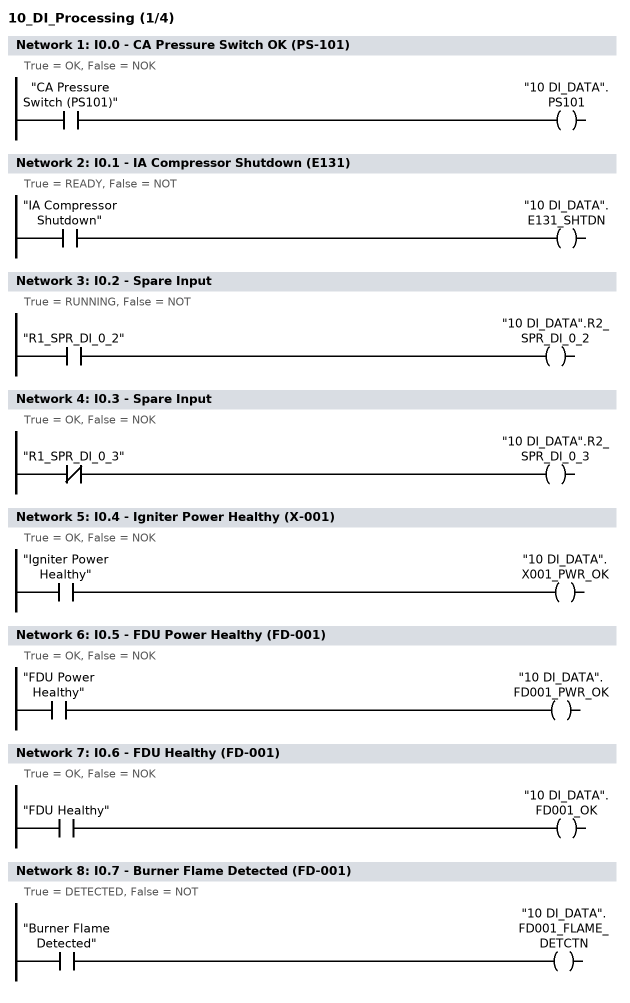
   RUNG wire#powerrail
      Contact( "CA Pressure Switch (PS101)" )
      Coil( "10 DI_DATA".PS101 )
   END_RUNG
   // the same network as SCL:
   "10 DI_DATA".PS101 := "CA Pressure Switch (PS101)";
END_REGION

REGION Network 2: I0.1 - IA Compressor Shutdown (E131)
   // True = READY, False = NOT
   RUNG wire#powerrail
      Contact( "IA Compressor Shutdown" )
      Coil( "10 DI_DATA".E131_SHTDN )
   END_RUNG
   // the same network as SCL:
   "10 DI_DATA".E131_SHTDN := "IA Compressor Shutdown";
END_REGION

REGION Network 3: I0.2 - Spare Input
   // True = RUNNING, False = NOT
   RUNG wire#powerrail
      Contact( "R1_SPR_DI_0_2" )
      Coil( "10 DI_DATA".R2_SPR_DI_0_2 )
   END_RUNG
   // the same network as SCL:
   "10 DI_DATA".R2_SPR_DI_0_2 := "R1_SPR_DI_0_2";
END_REGION

REGION Network 4: I0.3 - Spare Input
   // True = OK, False = NOK
   RUNG wire#powerrail
      I_Contact( "R1_SPR_DI_0_3" )
      Coil( "10 DI_DATA".R2_SPR_DI_0_3 )
   END_RUNG
   // the same network as SCL:
   "10 DI_DATA".R2_SPR_DI_0_3 := NOT "R1_SPR_DI_0_3";
END_REGION

REGION Network 5: I0.4 - Igniter Power Healthy (X-001)
   // True = OK, False = NOK
   RUNG wire#powerrail
      Contact( "Igniter Power Healthy" )
      Coil( "10 DI_DATA".X001_PWR_OK )
   END_RUNG
   // the same network as SCL:
   "10 DI_DATA".X001_PWR_OK := "Igniter Power Healthy";
END_REGION

REGION Network 6: I0.5 - FDU Power Healthy (FD-001)
   // True = OK, False = NOK
   RUNG wire#powerrail
      Contact( "FDU Power Healthy" )
      Coil( "10 DI_DATA".FD001_PWR_OK )
   END_RUNG
   // the same network as SCL:
   "10 DI_DATA".FD001_PWR_OK := "FDU Power Healthy";
END_REGION

REGION Network 7: I0.6 - FDU Healthy (FD-001)
   // True = OK, False = NOK
   RUNG wire#powerrail
      Contact( "FDU Healthy" )
      Coil( "10 DI_DATA".FD001_OK )
   END_RUNG
   // the same network as SCL:
   "10 DI_DATA".FD001_OK := "FDU Healthy";
END_REGION

REGION Network 8: I0.7 - Burner Flame Detected (FD-001)
   // True = DETECTED, False = NOT
   RUNG wire#powerrail
      Contact( "Burner Flame Detected" )
      Coil( "10 DI_DATA".FD001_FLAME_DETCTN )
   END_RUNG
   // the same network as SCL:
   "10 DI_DATA".FD001_FLAME_DETCTN := "Burner Flame Detected";
END_REGION

REGION Network 9: I1.0 - Pilot Ignition Air Flow Switch (FS-123)
   // True = FLOW, False = NO FLOW
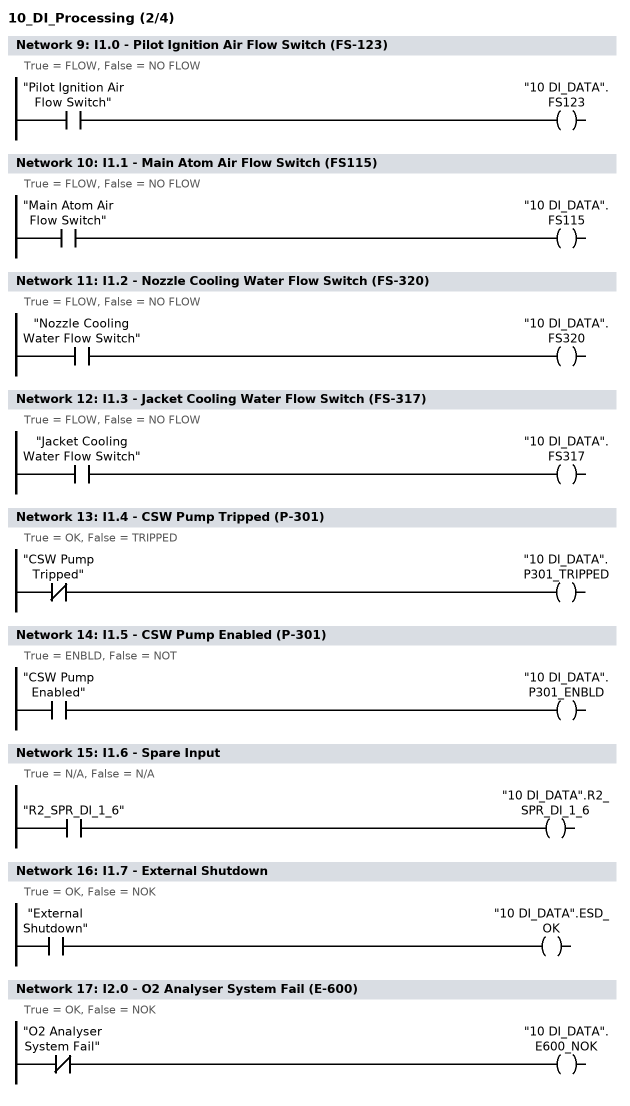
   RUNG wire#powerrail
      Contact( "Pilot Ignition Air Flow Switch" )
      Coil( "10 DI_DATA".FS123 )
   END_RUNG
   // the same network as SCL:
   "10 DI_DATA".FS123 := "Pilot Ignition Air Flow Switch";
END_REGION

REGION Network 10: I1.1 - Main Atom Air Flow Switch (FS115)
   // True = FLOW, False = NO FLOW
   RUNG wire#powerrail
      Contact( "Main Atom Air Flow Switch" )
      Coil( "10 DI_DATA".FS115 )
   END_RUNG
   // the same network as SCL:
   "10 DI_DATA".FS115 := "Main Atom Air Flow Switch";
END_REGION

REGION Network 11: I1.2 - Nozzle Cooling Water Flow Switch (FS-320)
   // True = FLOW, False = NO FLOW
   RUNG wire#powerrail
      Contact( "Nozzle Cooling Water Flow Switch" )
      Coil( "10 DI_DATA".FS320 )
   END_RUNG
   // the same network as SCL:
   "10 DI_DATA".FS320 := "Nozzle Cooling Water Flow Switch";
END_REGION

REGION Network 12: I1.3 - Jacket Cooling Water Flow Switch (FS-317)
   // True = FLOW, False = NO FLOW
   RUNG wire#powerrail
      Contact( "Jacket Cooling Water Flow Switch" )
      Coil( "10 DI_DATA".FS317 )
   END_RUNG
   // the same network as SCL:
   "10 DI_DATA".FS317 := "Jacket Cooling Water Flow Switch";
END_REGION

REGION Network 13: I1.4 - CSW Pump Tripped (P-301)
   // True = OK, False = TRIPPED
   RUNG wire#powerrail
      I_Contact( "CSW Pump Tripped" )
      Coil( "10 DI_DATA".P301_TRIPPED )
   END_RUNG
   // the same network as SCL:
   "10 DI_DATA".P301_TRIPPED := NOT "CSW Pump Tripped";
END_REGION

REGION Network 14: I1.5 - CSW Pump Enabled (P-301)
   // True = ENBLD, False = NOT
   RUNG wire#powerrail
      Contact( "CSW Pump Enabled" )
      Coil( "10 DI_DATA".P301_ENBLD )
   END_RUNG
   // the same network as SCL:
   "10 DI_DATA".P301_ENBLD := "CSW Pump Enabled";
END_REGION

REGION Network 15: I1.6 - Spare Input
   // True = N/A, False = N/A
   RUNG wire#powerrail
      Contact( "R2_SPR_DI_1_6" )
      Coil( "10 DI_DATA".R2_SPR_DI_1_6 )
   END_RUNG
   // the same network as SCL:
   "10 DI_DATA".R2_SPR_DI_1_6 := "R2_SPR_DI_1_6";
END_REGION

REGION Network 16: I1.7 - External Shutdown
   // True = OK, False = NOK
   RUNG wire#powerrail
      Contact( "External Shutdown" )
      Coil( "10 DI_DATA".ESD_OK )
   END_RUNG
   // the same network as SCL:
   "10 DI_DATA".ESD_OK := "External Shutdown";
END_REGION

REGION Network 17: I2.0 - O2 Analyser System Fail (E-600)
   // True = OK, False = NOK
   RUNG wire#powerrail
      I_Contact( "O2 Analyser System Fail" )
      Coil( "10 DI_DATA".E600_NOK )
   END_RUNG
   // the same network as SCL:
   "10 DI_DATA".E600_NOK := NOT "O2 Analyser System Fail";
END_REGION

REGION Network 18: I2.1 - O2 Analyser HiHi (E-600)
   // True = OK, False = HIHI
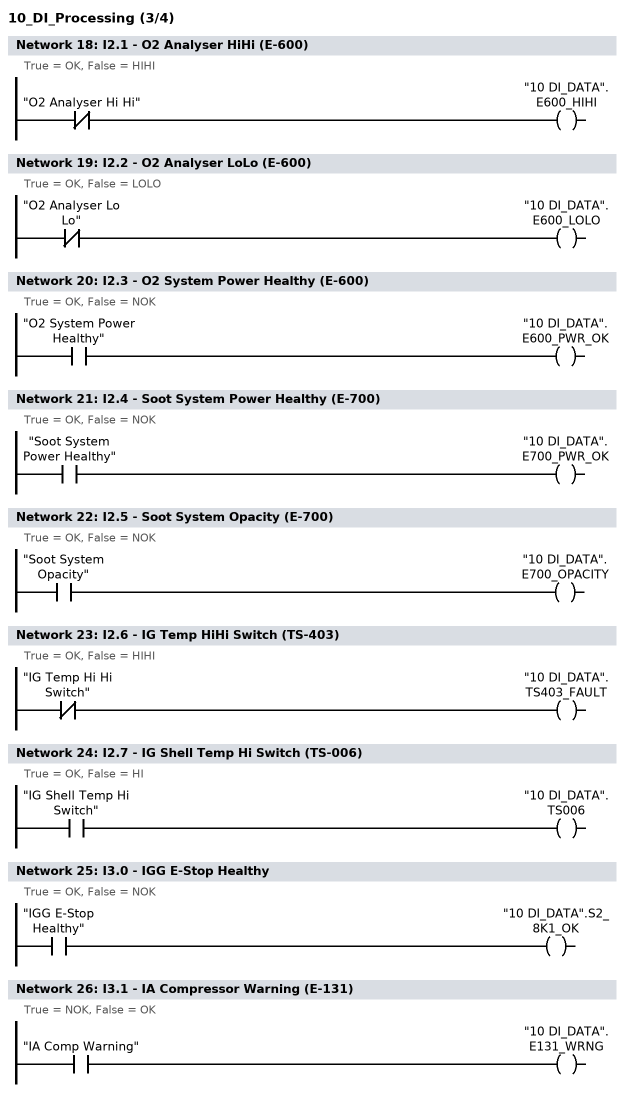
   RUNG wire#powerrail
      I_Contact( "O2 Analyser Hi Hi" )
      Coil( "10 DI_DATA".E600_HIHI )
   END_RUNG
   // the same network as SCL:
   "10 DI_DATA".E600_HIHI := NOT "O2 Analyser Hi Hi";
END_REGION

REGION Network 19: I2.2 - O2 Analyser LoLo (E-600)
   // True = OK, False = LOLO
   RUNG wire#powerrail
      I_Contact( "O2 Analyser Lo Lo" )
      Coil( "10 DI_DATA".E600_LOLO )
   END_RUNG
   // the same network as SCL:
   "10 DI_DATA".E600_LOLO := NOT "O2 Analyser Lo Lo";
END_REGION

REGION Network 20: I2.3 - O2 System Power Healthy (E-600)
   // True = OK, False = NOK
   RUNG wire#powerrail
      Contact( "O2 System Power Healthy" )
      Coil( "10 DI_DATA".E600_PWR_OK )
   END_RUNG
   // the same network as SCL:
   "10 DI_DATA".E600_PWR_OK := "O2 System Power Healthy";
END_REGION

REGION Network 21: I2.4 - Soot System Power Healthy (E-700)
   // True = OK, False = NOK
   RUNG wire#powerrail
      Contact( "Soot System Power Healthy" )
      Coil( "10 DI_DATA".E700_PWR_OK )
   END_RUNG
   // the same network as SCL:
   "10 DI_DATA".E700_PWR_OK := "Soot System Power Healthy";
END_REGION

REGION Network 22: I2.5 - Soot System Opacity (E-700)
   // True = OK, False = NOK
   RUNG wire#powerrail
      Contact( "Soot System Opacity" )
      Coil( "10 DI_DATA".E700_OPACITY )
   END_RUNG
   // the same network as SCL:
   "10 DI_DATA".E700_OPACITY := "Soot System Opacity";
END_REGION

REGION Network 23: I2.6 - IG Temp HiHi Switch (TS-403)
   // True = OK, False = HIHI
   RUNG wire#powerrail
      I_Contact( "IG Temp Hi Hi Switch" )
      Coil( "10 DI_DATA".TS403_FAULT )
   END_RUNG
   // the same network as SCL:
   "10 DI_DATA".TS403_FAULT := NOT "IG Temp Hi Hi Switch";
END_REGION

REGION Network 24: I2.7 - IG Shell Temp Hi Switch (TS-006)
   // True = OK, False = HI
   RUNG wire#powerrail
      Contact( "IG Shell Temp Hi Switch" )
      Coil( "10 DI_DATA".TS006 )
   END_RUNG
   // the same network as SCL:
   "10 DI_DATA".TS006 := "IG Shell Temp Hi Switch";
END_REGION

REGION Network 25: I3.0 - IGG E-Stop Healthy
   // True = OK, False = NOK
   RUNG wire#powerrail
      Contact( "IGG E-Stop Healthy" )
      Coil( "10 DI_DATA".S2_8K1_OK )
   END_RUNG
   // the same network as SCL:
   "10 DI_DATA".S2_8K1_OK := "IGG E-Stop Healthy";
END_REGION

REGION Network 26: I3.1 - IA Compressor Warning (E-131)
   // True = NOK, False = OK
   RUNG wire#powerrail
      Contact( "IA Comp Warning" )
      Coil( "10 DI_DATA".E131_WRNG )
   END_RUNG
   // the same network as SCL:
   "10 DI_DATA".E131_WRNG := "IA Comp Warning";
END_REGION

